   REGION "PAGE UP"
       //#hmi.page_up_actuate := #plc.pageUp.actuate;
       #hmi.page_up_animate := #plc.pageUp.animate;
       #hmi.page_up_enable := #plc.pageUp.enable;
       #hmi.page_up_label := #plc.pageUp.label;
       #hmi.page_up_list_select := #plc.pageUp.listSelect;
       #hmi.page_up_visible := #plc.pageUp.visible;
   END_REGION


   REGION "LINE UP"
       //#hmi.line_up_actuate := #plc.lineUp.actuate;
       #hmi.line_up_animate := #plc.lineUp.animate;
       #hmi.line_up_enable := #plc.lineUp.enable;
       #hmi.line_up_label := #plc.lineUp.label;
       #hmi.line_up_list_select := #plc.lineUp.listSelect;
       #hmi.line_up_visible := #plc.lineUp.visible;
   END_REGION


   REGION "LINE DOWN"
       //#hmi.line_down_actuate := #plc.lineDown.actuate;
       #hmi.line_down_animate := #plc.lineDown.animate;
       #hmi.line_down_enable := #plc.lineDown.enable;
       #hmi.line_down_label := #plc.lineDown.label;
       #hmi.line_down_list_select := #plc.lineDown.listSelect;
       #hmi.line_down_visible := #plc.lineDown.visible;
   END_REGION


   REGION "PAGE DOWN"
       //#hmi.page_down_actuate := #plc.pageDown.actuate;
       #hmi.page_down_animate := #plc.pageDown.animate;
       #hmi.page_down_enable := #plc.pageDown.enable;
       #hmi.page_down_label := #plc.pageDown.label;
       #hmi.page_down_list_select := #plc.pageDown.listSelect;
       #hmi.page_down_visible := #plc.pageDown.visible;
   END_REGION

   REGION "BOTTOM"
       //#hmi.bottom_actuate := #plc.bottom.actuate;
       #hmi.bottom_animate := #plc.bottom.animate;
       #hmi.bottom_enable := #plc.bottom.enable;
       #hmi.bottom_label := #plc.bottom.label;
       #hmi.bottom_list_select := #plc.bottom.listSelect;
       #hmi.bottom_visible := #plc.bottom.visible;
   END_REGION
END_FUNCTION

FUNCTION "NavBar: Private: First Row" : DInt   // FC180, SCL
{ S7_Optimized_Access := 'TRUE' }
VERSION : 0.1
   VAR_INPUT
      first_row : DInt;
      offset : DInt;
      TABLE_LENGTH : DInt;
   END_VAR
   VAR_TEMP
      ret : DInt;
   END_VAR
BEGIN
   REGION "DESCRIPTION"
       (*
       The new first row of the table is calculated from the offset. 
       Rollover and rollunder are resolved for the first row.
       *)
   END_REGION

   REGION "COPY TO INTERNAL"
       #ret := #first_row + #offset;
   END_REGION

   REGION "ROLLUNDER"
       IF #ret < 0 THEN
           #ret := #ret + #TABLE_LENGTH + 1;
       END_IF;
   END_REGION

   REGION "ROLLOVER"
       IF #ret > #TABLE_LENGTH THEN
           #ret := #ret - #TABLE_LENGTH - 1;
       END_IF;
   END_REGION

   REGION "OUTPUT"
       #"NavBar: Private: First Row" := #ret;
   END_REGION
END_FUNCTION

// folder: Utilities/Part Number

FUNCTION_BLOCK "IO Field: State Changes"   // FB48, SCL
{ S7_Optimized_Access := 'TRUE' }
VERSION : 0.1
   VAR_IN_OUT
      interface : "IO Field Data: Label with Data";
      feedback : "IO Field: State Change Data";
   END_VAR
   VAR
      old : "IO Field Data: Label with Data";
   END_VAR
BEGIN
   REGION "ANIMATE"
       #feedback.animate.rising := "USInt.Value_Change"(value := #interface.animate,
                                                         old_value := #old.animate);
       #feedback.animate.actual := #interface.animate;
       #feedback.animate.falling := FALSE;     // animate never set to null token 
   END_REGION

   REGION "ENABLE"
       #feedback.enable.rising := "Bool.Rising_Edge"(signal := #interface.enable,
                                                      old_signal := #old.enable);
       #feedback.enable.actual := #interface.enable;
       #feedback.enable.falling := "Bool.Falling_Edge"(signal := #interface.enable,
                                                        old_signal := #old.enable);
   END_REGION

   REGION "INPUT FINISHED"
       #feedback.input_finished.rising := "Bool.Rising_Edge"(signal := #interface.input_finished,
                                                              old_signal := #old.input_finished);
       #feedback.input_finished.actual := #interface.input_finished;
       #feedback.input_finished.falling := "Bool.Falling_Edge"(signal := #interface.input_finished,
                                                                old_signal := #old.input_finished);
   END_REGION

   REGION "VALUE CHANGED"
       #feedback.value.rising := "WString.Rising_Edge"(value := #interface.value,
                                                        old_value := #old.value);
       #feedback.value.actual := #interface.value;
       #feedback.value.falling := "WString.Falling_Edge"(value := #interface.value,
                                                          old_value := #old.value);
   END_REGION

   REGION "VISIBLE"
       #feedback.visible.rising := "Bool.Rising_Edge"(signal := #interface.visible,
                                                       old_signal := #old.visible);
       #feedback.visible.actual := #interface.visible;
       #feedback.visible.falling := "Bool.Falling_Edge"(signal := #interface.visible,
                                                         old_signal := #old.visible);
   END_REGION

   REGION "SAVE OLD VALUES"
       #old := #interface;
   END_REGION
END_FUNCTION_BLOCK

FUNCTION "Part_Number.Parse_Code" : Void   // FC34, SCL
{ S7_Optimized_Access := 'TRUE' }
VERSION : 0.1
   VAR_INPUT
      code : DInt;
   END_VAR
   VAR_OUTPUT
      code_left : DInt;
      code_right : DInt;
   END_VAR
BEGIN
   IF #code > 0 THEN
       #code_left := #code / 1000;
       #code_right := #code - #code / 1000 * 1000;
   ELSE
       #code_left := 0;
       #code_right := 0;
   END_IF;
END_FUNCTION

FUNCTION "Part_Number.Code_to_WString" : WString   // FC37, SCL
{ S7_Optimized_Access := 'TRUE' }
VERSION : 0.1
   VAR_INPUT
      pnLib : "Recipe: PN Text Library";
      pnCode : DInt;
   END_VAR
   VAR_TEMP
      pnLeft : DInt;
      pnRight : DInt;
      output : WString;
   END_VAR
   VAR CONSTANT
      newLine : WString := WSTRING#'$L';
   END_VAR
BEGIN
   REGION "PARSE CODE"
       "Part_Number.Parse_Code"(code := #pnCode,
                                 code_left => #pnLeft,
                                 code_right => #pnRight);
   END_REGION

   REGION "SINGLE LINE PN"
       IF "Part_Number.Is_Single"(#pnCode) THEN
           #output := #pnLib.pnText[#pnLeft];
       END_IF;
   END_REGION

   REGION "DOUBLE LINE PN"
       IF "Part_Number.Is_Double"(#pnCode) THEN
           #output := CONCAT_WSTRING(IN1 := #pnLib.pnText[#pnLeft],
                                     IN2 := #newLine,
                                     IN3 := #pnLib.pnText[#pnRight]);
       END_IF;
   END_REGION

   REGION "OUTPUT"
       #"Part_Number.Code_to_WString" := #output;
   END_REGION
END_FUNCTION

FUNCTION "Part_Number.Is_Double" : Bool   // FC153, SCL
{ S7_Optimized_Access := 'TRUE' }
VERSION : 0.1
   VAR_INPUT
      code : DInt;
   END_VAR
   VAR_TEMP
      code_left : DInt;
      code_right : DInt;
      ret : Bool;
   END_VAR
BEGIN
   REGION "NOTES"
       (*
       Double codes have a non-zero right hand component.
       Structure: XXXYYY
       XXX: left code, used for single and double codes
       YYY: right code, only used for double codes
       Last Edit: 2021-10-07
       *)
   END_REGION

   REGION "PROCESS CODE"
       "Part_Number.Parse_Code"(code := #code,
                                code_left => #code_left,
                                code_right => #code_right);
   END_REGION

   REGION "CHECK FOR DOUBLE CODE"
       IF #code_right > 0 THEN
           #ret := TRUE;
       END_IF;
   END_REGION

   REGION "RETURN" 
       #"Part_Number.Is_Double" := #ret;
   END_REGION
END_FUNCTION

FUNCTION "Part_Number.Is_Single" : Bool   // FC154, SCL
{ S7_Optimized_Access := 'TRUE' }
VERSION : 0.1
   VAR_INPUT
      code : DInt;
   END_VAR
   VAR_TEMP
      code_left : DInt;
      code_right : DInt;
      ret : Bool;
   END_VAR
BEGIN
   REGION "NOTES"
       (*
       Double codes have a non-zero right hand component.
       Structure:
       XXXYYY
       XXX: left code, used for single and double codes
       YYY: right code, only used for double codes
       Last Edit: 2021-10-07
       *)
   END_REGION

   REGION "PROCESS CODE"
       "Part_Number.Parse_Code"(code := #code,
                                code_left => #code_left,
                                code_right => #code_right);
   END_REGION

   REGION "CHECK FOR DOUBLE CODE"
       IF #code_right = 0 THEN
           #ret := TRUE;
       END_IF;
   END_REGION

   REGION "RETURN" 
       #"Part_Number.Is_Single" := #ret;
   END_REGION
END_FUNCTION

FUNCTION "Part_Number.WString_to_Code" : DInt   // FC240, SCL
{ S7_Optimized_Access := 'TRUE' }
VERSION : 0.1
   VAR_INPUT
      part_number : WString;
   END_VAR
   VAR_IN_OUT
      pn_library : "Recipe: PN Text Library";
   END_VAR
   VAR_TEMP
      _in_library : Bool;
      _library_full : Bool;
      _part_numbers : Array[0..1] of WString;
      _partial_pn_code : DInt;
      _pn_count : Int;
      _pn_code : DInt;
   END_VAR
   VAR CONSTANT
      OUT_OF_MEMORY : DInt := 999;
   END_VAR
BEGIN
   REGION "DATA PREP""
       "Part_Number.Split_PNs"(part_number := #part_number,
                               part_numbers := #_part_numbers);
       #_pn_count := "Part_Number.Count_PNs"(#_part_numbers);
   END_REGION


   REGION "NO PART NUMBERS ENTERED"
       IF #_pn_count = 0 THEN
           #"Part_Number.WString_to_Code" := 0;
           RETURN;
       END_IF;
   END_REGION


   REGION "CHECK FIRST PN CODE"
       #_pn_code := "Part_Number_Library.Search"(pn_library := #pn_library,
                                                 search_term := #_part_numbers[0]);
       #_in_library := "Part_Number.In_Library"(#_pn_code);
       #_library_full := "Part_Number_Library.Is_Full"(#pn_library);
   END_REGION


   REGION "FIRST PN CODE IN LIBRARY"
       IF #_in_library THEN
           #_pn_code *= 1_000;
       END_IF;
   END_REGION


   REGION "FIRST PN NOT IN LIBRARY, NO SPACE"
       IF NOT #_in_library AND #_library_full THEN
           #_pn_code := #OUT_OF_MEMORY * 1_000;
       END_IF;
   END_REGION


   REGION "FIRST PN NOT IN LIBRARY, SPACE"
       IF NOT #_in_library AND NOT #_library_full THEN
           #_pn_code := 1_000 * "Part_Number_Library.Add_PN"(pn := #_part_numbers[0],
                                                             pn_library := #pn_library);
       END_IF;
   END_REGION


   REGION "RETURN SINGLE PN CODE"
       IF #_pn_count = 1 THEN
           #"Part_Number.WString_to_Code" := #_pn_code;
           RETURN;
       END_IF;
   END_REGION


   REGION "CHECK SECOND PN CODE"
       #_partial_pn_code := "Part_Number_Library.Search"(pn_library := #pn_library,
                                                         search_term := #_part_numbers[1]);
       #_in_library := "Part_Number.In_Library"(#_partial_pn_code);
       #_library_full := "Part_Number_Library.Is_Full"(#pn_library);
   END_REGION


   REGION "SECOND PN CODE IN LIBRARY"
       IF #_in_library THEN
           #"Part_Number.WString_to_Code" := #_pn_code + #_partial_pn_code;
           RETURN;
       END_IF;
   END_REGION


   REGION "SECOND PN NOT IN LIBRARY, NO SPACE"
       IF NOT #_in_library AND #_library_full THEN
           #"Part_Number.WString_to_Code" := #_pn_code + #OUT_OF_MEMORY;
           RETURN;
       END_IF;
   END_REGION


   REGION "SECOND PN NOT IN LIBRARY, SPACE"
       IF NOT #_in_library AND NOT #_library_full THEN
           #_pn_code += "Part_Number_Library.Add_PN"(pn := #_part_numbers[1],
                                                     pn_library := #pn_library);
           #"Part_Number.WString_to_Code" := #_pn_code;
           RETURN;
       END_IF;
   END_REGION


   #"Part_Number.WString_to_Code" := 0;
   RETURN;
END_FUNCTION

FUNCTION "Part_Number.Count_PNs" : Int   // FC252, SCL
{ S7_Optimized_Access := 'TRUE' }
VERSION : 0.1
   VAR_INPUT
      part_numbers : Array[0..1] of WString;
   END_VAR
   VAR CONSTANT
      NULL : WString := WSTRING#'//';
      BLANK : WString := WSTRING#'';
   END_VAR
BEGIN
   IF #part_numbers[0] = #NULL THEN
       #"Part_Number.Count_PNs" := 0;
       RETURN;
   END_IF;

   IF #part_numbers[0] = #BLANK THEN
       #"Part_Number.Count_PNs" := 0;
       RETURN;
   END_IF;

   IF #part_numbers[1] = #NULL THEN
       #"Part_Number.Count_PNs" := 1;
       RETURN;
   END_IF;

   IF #part_numbers[1] = #BLANK THEN
       #"Part_Number.Count_PNs" := 1;
       RETURN;
   END_IF;

   #"Part_Number.Count_PNs" := 2;
   RETURN;
END_FUNCTION

FUNCTION "Part_Number.In_Library" : Bool   // FC253, SCL
{ S7_Optimized_Access := 'TRUE' }
VERSION : 0.1
   VAR_INPUT
      pn_code : DInt;
   END_VAR
BEGIN
   IF #pn_code = "NULL_TOKEN" THEN
       #"Part_Number.In_Library" := FALSE;
       RETURN;
   END_IF;
   #"Part_Number.In_Library" := TRUE;
   RETURN;
END_FUNCTION

FUNCTION "Part_Number.Split_PNs" : Void   // FC254, SCL
{ S7_Optimized_Access := 'TRUE' }
VERSION : 0.1
   VAR_INPUT
      part_number : WString;
   END_VAR
   VAR_IN_OUT
      part_numbers : Array[0..1] of WString;
   END_VAR
   VAR_TEMP
      _part_numbers : Array[0..1] of WString;
   END_VAR
   VAR CONSTANT
      NEW_LINE : WString := WSTRING#'$L';
      NULL : WString := WSTRING#'//';
   END_VAR
BEGIN
   "Array.WString.Fill"(value := #NULL,
                        array := #_part_numbers);
   "WString.Split_Single"(wstring_in := #part_number,
                          delimeter := #NEW_LINE,
                          "pointer" := 0,
                          sub_strings := #_part_numbers);
   #part_numbers := #_part_numbers;
END_FUNCTION

// folder: Utilities/Part Number Library

FUNCTION "Part_Number_Library.Is_Full" : Bool   // FC250, SCL
{ S7_Optimized_Access := 'TRUE' }
VERSION : 0.1
   VAR_INPUT
      pn_library : "Recipe: PN Text Library";
   END_VAR
   VAR_TEMP
      _first_null : DInt;
   END_VAR
   VAR CONSTANT
      NULL_STRING : WString := WSTRING#'//';
   END_VAR
BEGIN
   #_first_null := "Part_Number_Library.Search"(pn_library := #pn_library,
                                                search_term := #NULL_STRING);
   IF #_first_null = "NULL_TOKEN" THEN
       #"Part_Number_Library.Is_Full" := TRUE;
       RETURN;
   END_IF;

   #"Part_Number_Library.Is_Full" := FALSE;
   RETURN;
END_FUNCTION

FUNCTION "Part_Number_Library.Add_PN" : DInt   // FC251, SCL
{ S7_Optimized_Access := 'TRUE' }
VERSION : 0.1
   VAR_INPUT
      pn : WString;
   END_VAR
   VAR_IN_OUT
      pn_library : "Recipe: PN Text Library";
   END_VAR
   VAR_TEMP
      _index : DInt;
   END_VAR
   VAR CONSTANT
      NULL_STRING : WString := WSTRING#'//';
   END_VAR
BEGIN
   #_index := "Part_Number_Library.Search"(pn_library := #pn_library,
                                           search_term := #NULL_STRING);
   #pn_library.pnText[#_index] := #pn;
   #"Part_Number_Library.Add_PN" := #_index;
END_FUNCTION

FUNCTION "Part_Number_Library.Search" : Int   // FC255, SCL
{ S7_Optimized_Access := 'TRUE' }
VERSION : 0.1
   VAR_INPUT
      pn_library : "Recipe: PN Text Library";
      search_term : WString;
   END_VAR
   VAR_TEMP
      _array : Array[0..#MAX_ELEMENTS] of WString;
      _slices : Int;
      _slice : Int;
      _internal_length : Int;
      _external_length : Int;
      _search_result : Int;
   END_VAR
   VAR CONSTANT
      MAX_ELEMENTS : Int := 24;
   END_VAR
BEGIN
   REGION "NOTES"
       (*
           Why is this necessary?
               Unfortunately, dynamically sized arrays of wstring data type cannot accept
               wstrings of a declared length (e.x. the input parameter array[*] of 
               wstring[10] cannot exist). We need this wrapper function so that we can 
               copy wstrings of a declared length to an array of wstrings of default 
               length. Once copied, this array can be passed into the wstring search 
               function. However, there is only 16k of local memory to store the array of
               wstrings of default length. The pn text library can store up to 1000 part 
               numbers. If we were to copy all 1000, we would need 500k of memory. So, we 
               must slice the pn library into chunks and search them.
           Why are part number text wstrings a declared length?
               The declared lenght was necessary to fit a reasonable number of part 
               numbers into retentive memory.
       *)
   END_REGION


   REGION "SETUP"
       #_internal_length := UDINT_TO_INT("Array.Any.Length"(#_array));
       #_external_length := UDINT_TO_INT("Array.Any.Length"(#pn_library.pnText));
       #_slices := #_external_length / #_internal_length - 1;
   END_REGION


   REGION "REPEAT FOR EACH SLICE OF EXTERNAL ARRAY"
       FOR #_slice := 0 TO #_slices DO
           "Part_Number_Library.Search.Map_to_Internal_Array"(pn_library := #pn_library,
                                                              slice_number := #_slice,
                                                              internal_array := #_array);
           #_search_result := "Array.WString.Search"(array := #_array,
                                                     search_term := #search_term);
           IF #_search_result <> "NULL_TOKEN" THEN
               #"Part_Number_Library.Search" := #_search_result + #_slice * #_internal_length;
               RETURN;
           END_IF;
       END_FOR;
   END_REGION

   REGION "RETURN"
       #"Part_Number_Library.Search" := "NULL_TOKEN";
       RETURN;
   END_REGION
END_FUNCTION

FUNCTION "Part_Number_Library.Search.Map_to_Internal_Array" : Void   // FC256, SCL
{ S7_Optimized_Access := 'TRUE' }
VERSION : 0.1
   VAR_INPUT
      pn_library : "Recipe: PN Text Library";
      slice_number : Int;
   END_VAR
   VAR_IN_OUT
      internal_array : Array[*] of WString;
   END_VAR
   VAR_TEMP
      _i : Int;
      _length : Int;
      _p : Int;
   END_VAR
BEGIN
   #_length := UDINT_TO_INT("Array.Any.Length"(#internal_array));
   FOR #_i := 0 TO #_length - 1 DO
       #_p := #_i + #slice_number * #_length;
       #internal_array[#_i] := #pn_library.pnText[#_p];
   END_FOR;
END_FUNCTION

// folder: Utilities/Real

FUNCTION_BLOCK "Real.State_Change"   // FB52, SCL
{ S7_Optimized_Access := 'TRUE' }
VERSION : 0.1
   VAR_INPUT
      value : Real;
   END_VAR
   VAR_IN_OUT
      get_real : "State Changes: Real";
   END_VAR
   VAR
      old_value : Real;
   END_VAR
   VAR_TEMP
      _return : "State Changes: Real";
   END_VAR
BEGIN
   REGION "BUFFER IN"
       #_return := #get_real;
   END_REGION

   REGION "MAP"
       IF #value <> #old_value THEN
           #_return.actual := #value;
       END_IF;
       // these are set to false because there are no invalid times
       // negative should count in reverse
       // zero is valid
       #_return.rising := FALSE;
       #_return.falling := FALSE;
   END_REGION

   REGION "SAVE OLD VALUE"
       #old_value := #value;
   END_REGION


   REGION "RETURN" 
       #get_real := #_return;
   END_REGION
END_FUNCTION_BLOCK

// folder: Utilities/Screen Objects

FUNCTION "Cell_Data.Hide" : "Cell Data"   // FC209, SCL
{ S7_Optimized_Access := 'TRUE' }
VERSION : 0.1
BEGIN
   #"Cell_Data.Hide".animate := "INVISIBLE";
   #"Cell_Data.Hide".data := "BLANK";
   #"Cell_Data.Hide".visibility := "HIDE";
END_FUNCTION

FUNCTION "Cell_Data.Show" : "Cell Data"   // FC216, SCL
{ S7_Optimized_Access := 'TRUE' }
VERSION : 0.1
   VAR_INPUT
      animate : Int;
      data : WString;
   END_VAR
   VAR_TEMP
      _ret : "Cell Data";
   END_VAR
BEGIN
   #_ret.animate := #animate;
   #_ret.data := #data;
   #_ret.visibility := "SHOW";
   #"Cell_Data.Show" := #_ret;
END_FUNCTION

// folder: Utilities/Selected Buttons

FUNCTION "Selected_Buttons.Indices" : Void   // FC246, SCL
{ S7_Optimized_Access := 'TRUE' }
VERSION : 0.1
   VAR_INPUT
      selected_buttons : "Selected Buttons";
   END_VAR
   VAR_IN_OUT
      selected_buttons_indices : Array[*] of Int;
   END_VAR
   VAR_TEMP
      _i : Int;
      _length : Int;
      _resized_bool_array : Array[0..999] of Bool;
   END_VAR
BEGIN
   "Array.Bool.True_Indices"(array_of_bool := #selected_buttons.btns,
                             length := "BUTTON_COUNT",
                             list_of_indices := #selected_buttons_indices);
   FOR #_i := 0 TO "BUTTON_COUNT" DO
       IF #selected_buttons_indices[#_i] = "NULL_TOKEN" THEN
           CONTINUE;
       END_IF;
       #selected_buttons_indices[#_i] := "KP8.DURL_to_LRUD"(#selected_buttons_indices[#_i]);
   END_FOR;
END_FUNCTION

FUNCTION "Selected_Buttons.Get_First_Selected_Button" : Int   // FC289, SCL
{ S7_Optimized_Access := 'TRUE' }
VERSION : 0.1
   VAR_INPUT
      selected_buttons : "Selected Buttons";
   END_VAR
   VAR_TEMP
      _selected_buttons : Array[0.."BUTTON_COUNT"] of Int;
   END_VAR
BEGIN
   "Selected_Buttons.Indices"(selected_buttons := #selected_buttons,
                              selected_buttons_indices := #_selected_buttons);
   #"Selected_Buttons.Get_First_Selected_Button" := #_selected_buttons[0];
END_FUNCTION

// folder: Utilities/Selected Stations

FUNCTION "Selected_Stations.Indices" : Void   // FC245, SCL
{ S7_Optimized_Access := 'TRUE' }
VERSION : 0.1
   VAR_INPUT
      selected_stations : "Selected Stations";
   END_VAR
   VAR_IN_OUT
      selected_stations_indices : Array[*] of Int;
   END_VAR
   VAR_TEMP
      _i : Int;
      _length : Int;
      _resized_array : Array[0..999] of Bool;
   END_VAR
BEGIN
   FOR #_i := 0 TO "STATION_COUNT" DO
       #_resized_array[#_i] := #selected_stations.stns[#_i];
   END_FOR;
   "Array.Bool.True_Indices"(array_of_bool := #_resized_array,
                             length := "STATION_COUNT",
                             list_of_indices := #selected_stations_indices);
END_FUNCTION

FUNCTION "Selected_Stations.Matching_Line_Names" : Bool   // FC257, SCL
{ S7_Optimized_Access := 'TRUE' }
VERSION : 0.1
   VAR_INPUT
      stations : "Station: All Stations";
      selected_stations : "Selected Stations";
   END_VAR
   VAR_TEMP
      _i : Int;
      _first_selected_line_name : WString;
   END_VAR
   // Ret_Val : returns true when any number of stations selected and all selected stations have matching names
   VAR CONSTANT
      BLANK : WString;
   END_VAR
BEGIN
   REGION "NOTES"
       (*
           2022-04-06
           returns true if all selected stations have matching names
           returns false if no station selected
           returns false if selected stations do not have matching names
       *)
   END_REGION


   REGION "RETURN FALSE IF NO STATIONS SELECTED"
       IF #selected_stations.count = 0 THEN
           #"Selected_Stations.Matching_Line_Names" := FALSE;
           RETURN;
       END_IF;
   END_REGION


   REGION "CHECK EACH STATION"
       FOR #_i := 0 TO "STATION_COUNT" DO

           REGION "IGNORE DE-SELECTED STATIONS"
               IF NOT #selected_stations.stns[#_i] THEN
                   CONTINUE;
               END_IF;
           END_REGION

           REGION "SAVE FIRST SELECTED STATION'S NAME"
               IF #_first_selected_line_name = #BLANK THEN
                   #_first_selected_line_name := #stations.stn[#_i].id.lineName;
                   CONTINUE;
               END_IF;
           END_REGION

           REGION "RETURN FALSE IF SELECTED STATIONS' NAMES DO NOT MATCH"
               IF #_first_selected_line_name <> #stations.stn[#_i].id.lineName THEN
                   #"Selected_Stations.Matching_Line_Names" := FALSE;
                   RETURN;
               END_IF;
           END_REGION

       END_FOR;
   END_REGION


   REGION "ALL SELECTED STATIONS HAVE MATCHING NAMES"
       #"Selected_Stations.Matching_Line_Names" := TRUE;
   END_REGION
END_FUNCTION

FUNCTION "Selected_Stations.Get_First_Selected_Station" : Int   // FC274, SCL
{ S7_Optimized_Access := 'TRUE' }
VERSION : 0.1
   VAR_INPUT
      selected_stations : "Selected Stations";
   END_VAR
   VAR_TEMP
      _selected_stations : Array[0.."STATION_COUNT"] of Int;
   END_VAR
BEGIN
   "Selected_Stations.Indices"(selected_stations := #selected_stations,
                               selected_stations_indices := #_selected_stations);
   #"Selected_Stations.Get_First_Selected_Station" := #_selected_stations[0];
END_FUNCTION

// folder: Utilities/String

FUNCTION "Strip Sign" : WString   // FC3, SCL
{ S7_Optimized_Access := 'TRUE' }
VERSION : 0.1
   VAR_INPUT
      WString : WString;
   END_VAR
   VAR_TEMP
      Length : Int;
      "String Box" : WString;
      "Test Character" : WString;
   END_VAR
   VAR CONSTANT
      "+" : WChar := WCHAR#'+';
      "-" : WChar := WCHAR#'-';
   END_VAR
BEGIN
   #"String Box" := #WString;
   #"Test Character" := LEFT_WSTRING(IN := #"String Box",
                                     L := 1);
   IF #"Test Character" = #"+" OR #"Test Character" = #"-" THEN
       #Length := LEN(#"String Box");
       #"String Box" := RIGHT_WSTRING(IN := #"String Box", L := #Length - 1);

   END_IF;
   #"Strip Sign" := #"String Box";
END_FUNCTION

FUNCTION "Add Leading" : WString   // FC4, SCL
{ S7_Optimized_Access := 'TRUE' }
VERSION : 0.1
   VAR_INPUT
      "Leading Character" : WChar;
      "Desired Length" : USInt;
      "String" : WString;
   END_VAR
   VAR_TEMP
      Length : Int;
      "String Box" : WString;
   END_VAR
BEGIN
   #"String Box" := #String;
   #Length := LEN(#"String Box");

   WHILE #Length < #"Desired Length" DO
       #"String Box" := CONCAT_WSTRING(IN1 := #"Leading Character",
                                       IN2 := #"String Box");
       #Length := LEN(#"String Box");
   END_WHILE;

   #"Add Leading" := #"String Box";
END_FUNCTION

FUNCTION "WString.Word_Wrap_Depricated" : WString   // FC28, SCL
{ S7_Optimized_Access := 'TRUE' }
VERSION : 0.1
   VAR_INPUT
      stringIn : WString;
      maxLength : Int;
   END_VAR
   VAR_TEMP
      length : Int;
      lineBox : Array[0..#limitLines] of WString["LONG_STRING_LENGTH"];
      ret : WString;
      stringBox : Array[0..#limitString] of WString["LONG_STRING_LENGTH"];
   END_VAR
   VAR CONSTANT
      space : WString := WSTRING#' ';
      blank : WString;
      lineBreak : WString := WSTRING#'$L';
      limitString : Int := 49;
      limitLines : Int := 9;
   END_VAR
BEGIN
   REGION "GET LENGTH"
       #length := LEN(#stringIn);
   END_REGION

   REGION "NO WRAP NECESSARY"
       IF #length <= #maxLength THEN
           #ret := #stringIn;
       END_IF;
   END_REGION


   REGION "EXECUTE WORD WRAP"
       IF #length > #maxLength THEN

           "Explode"(stringIn := #stringIn,
                     explodedString := #stringBox);

           "WString.Word_Wrap_Depricated.Construct_Line"(stringBox := #stringBox,
                                       lineBox := #lineBox,
                                       maxLength := #maxLength);

           #ret := "WString.Word_Wrap_Depricated.Concat_Lines"(#lineBox);

       END_IF;
   END_REGION

   REGION "RETURN"
       #"WString.Word_Wrap_Depricated" := #ret;
   END_REGION
END_FUNCTION

FUNCTION "Trim" : WString   // FC29, SCL
{ S7_Optimized_Access := 'TRUE' }
VERSION : 0.1
   VAR_INPUT
      wString : WString;
   END_VAR
   VAR_TEMP
      ret : WString;
   END_VAR
   VAR CONSTANT
      space : WString := WSTRING#' ';
   END_VAR
BEGIN
   #ret := #wString;
   WHILE LEFT(IN := #ret, L := 1) = #space DO
       #ret := RIGHT(IN := #ret, L := LEN(#ret) - 1);
   END_WHILE;
   WHILE RIGHT(IN := #ret, L := 1) = #space DO
       #ret := LEFT(IN := #ret, L := LEN(#ret) - 1);
   END_WHILE;
   #Trim := #ret;
END_FUNCTION

FUNCTION "Upper" : Void   // FC49, SCL
{ S7_Optimized_Access := 'TRUE' }
VERSION : 0.1
   VAR_IN_OUT
      "string" : Variant;
   END_VAR
   VAR_TEMP
      "type" : Bool;
      stringBox : String;
      status : Int;
      wStringBox : WString;
      charArr : Array[0..255] of Char;
      cntChar : UInt;
      pChar : Int;
   END_VAR
   VAR CONSTANT
      asciiLow : Char := 'a';
      asciiHigh : Char := 'z';
      asciiCaseOffset : Int := 32;
   END_VAR
BEGIN
   IF TypeOf(#string) = String THEN
       #status := MOVE_BLK_VARIANT(SRC := #string,
                                   COUNT := 1,
                                   SRC_INDEX := 0,
                                   DEST_INDEX := 0,
                                   DEST => #stringBox);
   ELSIF TypeOf(#string) = WString THEN
       #status := MOVE_BLK_VARIANT(SRC := #string,
                                   COUNT := 1,
                                   SRC_INDEX := 0,
                                   DEST_INDEX := 0,
                                   DEST => #wStringBox);
       #stringBox := WSTRING_TO_STRING(#wStringBox);
   ELSE
       RETURN;
   END_IF;

   Strg_TO_Chars(Strg := #stringBox,
                 pChars := 0,
                 Cnt => #cntChar,
                 Chars := #charArr);

   FOR #pChar := 0 TO UINT_TO_INT(#cntChar) - 1 DO
       IF #asciiLow <= #charArr[#pChar] AND #charArr[#pChar] <= #asciiHigh THEN
           #charArr[#pChar] := INT_TO_CHAR(CHAR_TO_INT(#charArr[#pChar]) - #asciiCaseOffset);
       END_IF;
   END_FOR;

   Chars_TO_Strg(Chars := #charArr,
                 pChars := 0,
                 Cnt := #cntChar,
                 Strg => #stringBox);

   IF TypeOf(#string) = String THEN
       #status := MOVE_BLK_VARIANT(SRC := #stringBox,
                                   COUNT := 1,
                                   SRC_INDEX := 0,
                                   DEST_INDEX := 0,
                                   DEST => #string);
   ELSIF TypeOf(#string) = WString THEN
       #wStringBox := STRING_TO_WSTRING(#stringBox);
       #status := MOVE_BLK_VARIANT(SRC := #wStringBox,
                                   COUNT := 1,
                                   SRC_INDEX := 0,
                                   DEST_INDEX := 0,
                                   DEST => #string);
   END_IF;
END_FUNCTION

FUNCTION "Explode" : Void   // FC73, SCL
{ S7_Optimized_Access := 'TRUE' }
VERSION : 0.1
   VAR_INPUT
      stringIn : WString;
   END_VAR
   VAR_IN_OUT
      explodedString : Variant;
   END_VAR
   VAR_TEMP
      charBox : Array[0..#lmtChar] of WChar;
      count : DInt;
      pChar : Int;
      pStringBox : Int;
      stringBox : Array[0..#lmtString] of WString["LONG_STRING_LENGTH"];
      status : DInt;
   END_VAR
   VAR CONSTANT
      space : WString := WSTRING#' ';
      blank : WString;
      lineBreak : WString := WSTRING#'$L';
      lmtString : Int := 49;
      lmtChar : Int := 999;
   END_VAR
BEGIN
   Strg_TO_Chars(Strg := #stringIn,
                 pChars := 0,
                 Cnt => #count,
                 Chars := #charBox);

   FOR #pChar := 0 TO #count DO

       IF #charBox[#pChar] = #space THEN
           IF #charBox[#pChar + 1] = #space THEN
               EXIT;
           END_IF;
       END_IF;

       IF #pChar = 0 THEN
           #stringBox[#pStringBox] := #charBox[#pChar];
       END_IF;

       IF #pChar >= 1 THEN
           #stringBox[#pStringBox] := CONCAT_WSTRING(IN1 := #stringBox[#pStringBox],
                                                     IN2 := #charBox[#pChar]);
       END_IF;

       IF #charBox[#pChar] = #space THEN
           #stringBox[#pStringBox] := "Trim"(#stringBox[#pStringBox]);
           #pStringBox := #pStringBox + 1;
       END_IF;

       IF #charBox[#pChar] = #lineBreak THEN
           #stringBox[#pStringBox] := LEFT(IN := #stringBox[#pStringBox],
                                           L := LEN(#stringBox[#pStringBox]) - 1);
           #pStringBox := #pStringBox + 1;
           #stringBox[#pStringBox] := #lineBreak;
           #pStringBox := #pStringBox + 1;
       END_IF;

   END_FOR;

   #status := MOVE_BLK_VARIANT(SRC := #stringBox,
                               COUNT := INT_TO_UDINT(#pStringBox)+1,
                               SRC_INDEX :=0,
                               DEST_INDEX := 0,
                               DEST => #explodedString);
END_FUNCTION

FUNCTION "WString.Word_Wrap_Depricated.Construct_Line" : Void   // FC74, SCL
{ S7_Optimized_Access := 'TRUE' }
VERSION : 0.1
   VAR_INPUT
      stringBox : Array[0..#limitString] of WString["LONG_STRING_LENGTH"];
      maxLength : Int;
   END_VAR
   VAR_IN_OUT
      lineBox : Array[0..#limitLines] of WString["LONG_STRING_LENGTH"];
   END_VAR
   VAR_TEMP
      _lineBox : Array[0..#limitLines] of WString["LONG_STRING_LENGTH"];
      pString : Int;
      pLineBox : Int;
      lengthTest : WString;
   END_VAR
   VAR CONSTANT
      space : WString := WSTRING#' ';
      blank : WString;
      lineBreak : WString := WSTRING#'$L';
      limitString : Int := 49;
      limitLines : Int := 9;
   END_VAR
BEGIN
   REGION "FOR EACH STRING IN STRING LIST"
       FOR #pString := 0 TO #limitString DO

           REGION "END OF STRING LIST"
               IF #stringBox[#pString] = #blank THEN
                   IF #stringBox[#pString + 1] = #blank THEN
                       #_lineBox[#pLineBox] := "Trim"(#_lineBox[#pLineBox]);
                       #lineBox := #_lineBox;
                       RETURN;
                   END_IF;
               END_IF;
           END_REGION

           REGION "ON NEW LINE CHARACTER"
               IF #stringBox[#pString] = #lineBreak THEN
                   #_lineBox[#pLineBox] := "Trim"(#_lineBox[#pLineBox]);
                   #pLineBox := #pLineBox + 1;
                   #_lineBox[#pLineBox] := #lineBreak;
                   #pLineBox := #pLineBox + 1;
               END_IF;
           END_REGION

           REGION "BUILD EACH LINE"
               IF #stringBox[#pString] <> #lineBreak THEN

                   REGION "FIRST ELEMENT EDGE CASE"
                       IF #pString = 0 THEN
                           #lengthTest := #stringBox[#pString];
                       END_IF;
                   END_REGION

                   REGION "BUILT TEST STRING"
                       IF #pString >= 1 THEN
                           #lengthTest := CONCAT_WSTRING(IN1 := #_lineBox[#pLineBox],
                                                         IN2 := #space,
                                                         IN3 := #stringBox[#pString]);
                       END_IF;
                   END_REGION

                   REGION "TEST STRING NOT TOO LONG"
                       IF LEN(#lengthTest) <= #maxLength THEN
                           #_lineBox[#pLineBox] := #lengthTest;
                       END_IF;
                   END_REGION

                   REGION "TEST STRING TOO LONG"
                       IF LEN(#lengthTest) > #maxLength THEN
                           #_lineBox[#pLineBox] := "Trim"(#_lineBox[#pLineBox]);
                           #_lineBox[#pLineBox] := "Trim"(#_lineBox[#pLineBox]);
                           #pLineBox := #pLineBox + 1;
                           #_lineBox[#pLineBox] := #stringBox[#pString];
                       END_IF;
                   END_REGION

               END_IF;
           END_REGION

       END_FOR;
   END_REGION

   REGION "RETURN"
       #lineBox := #_lineBox;
   END_REGION
END_FUNCTION

FUNCTION "WString.Word_Wrap_Depricated.Concat_Lines" : WString   // FC75, SCL
{ S7_Optimized_Access := 'TRUE' }
VERSION : 0.1
   VAR_INPUT
      lineBox : Array[0..#limitLines] of WString["LONG_STRING_LENGTH"];
   END_VAR
   VAR_TEMP
      pLine : Int;
      ret : WString;
   END_VAR
   VAR CONSTANT
      space : WString := WSTRING#' ';
      blank : WString;
      lineBreak : WString := WSTRING#'$L';
      limitString : Int := 49;
      limitLines : Int := 9;
   END_VAR
BEGIN
   REGION "FOR EACH LINE"
       FOR #pLine := 0 TO #limitLines DO

           REGION "ON END OF LINE LIST"
               IF #lineBox[#pLine] = #space OR #lineBox[#pLine] = #blank THEN
                   EXIT;
               END_IF;
           END_REGION

           REGION "ON FIRST ELEMENT IN LINE LIST"
               IF #pLine = 0 THEN
                   #ret := #lineBox[#pLine];
               END_IF;
           END_REGION

           REGION "CONSTRUCT OUTPUT"
               IF #pLine >= 1 THEN

                   REGION "NO OP ON LINE BREAK CHARACTER"
                       IF #lineBox[#pLine] = #lineBreak THEN
                           ;// no action required
                       END_IF;
                   END_REGION

                   REGION "CONCATINATION"
                       IF #lineBox[#pLine] <> #lineBreak THEN
                           #ret := CONCAT_WSTRING(IN1 := #ret,
                                                  IN2 := #lineBreak,
                                                  IN3 := #lineBox[#pLine]);
                       END_IF;
                   END_REGION

               END_IF;
           END_REGION


       END_FOR;
   END_REGION

   REGION "RETURN"
       #ret := "Trim"(#ret);
       #"WString.Word_Wrap_Depricated.Concat_Lines" := #ret;
   END_REGION
END_FUNCTION

FUNCTION "WString.Split_Single" : Void   // FC202, SCL
{ S7_Optimized_Access := 'TRUE' }
VERSION : 0.1
   VAR_INPUT
      wstring_in : WString;
      delimeter : WString;
      pointer : Int;
   END_VAR
   VAR_IN_OUT
      sub_strings : Array[*] of WString;
   END_VAR
   VAR_TEMP
      _split : WString;
      _position : Int;
      _return : WString;
   END_VAR
BEGIN
   REGION "GET POSITION OF DELIMETER IN STRING"
       #_position := FIND(IN1 := #wstring_in,
                          IN2 := #delimeter);
   END_REGION

   REGION "BASE CASE"
       IF #_position = 0 THEN
           #sub_strings[#pointer] := #wstring_in;
           RETURN;
       END_IF;
   END_REGION


   REGION "RECURSIVE CASE"
       #sub_strings[#pointer] := LEFT(IN := #wstring_in, L := #_position - 1);
       "WString.Split_Single"(wstring_in := RIGHT(IN := #wstring_in, L := LEN(#wstring_in) - #_position),
                       delimeter := #delimeter,
                       "pointer" := #pointer + 1,
                       sub_strings := #sub_strings);
   END_REGION
END_FUNCTION

FUNCTION "WString.Word_Wrap" : WString   // FC203, SCL
{ S7_Optimized_Access := 'TRUE' }
VERSION : 0.1
   VAR_INPUT
      delimeters : Array[*] of WString[1];
      line_length : Int;
      wstring_in : WString;
   END_VAR
   VAR_TEMP
      _i : Int;
      _substring_length : Int;
      _wstring_in_length : Int;
      _pointer_substrings : Int;
      _substring : WString;
      _position_of_last_delimeter : Int;
      _recurse : Bool;
      _string_split_right : WString;
   END_VAR
   VAR CONSTANT
      BLANK : WString;
      NEW_LINE : WString := WSTRING#'$L';
   END_VAR
BEGIN
   #_wstring_in_length := LEN(#wstring_in);

   IF #line_length = 0 THEN
       #"WString.Word_Wrap" := #BLANK;
       RETURN;
   END_IF;

   FOR #_i := 1 TO #_wstring_in_length DO

       #_substring := CONCAT_WSTRING(IN1 := #_substring,
                                     IN2 := #wstring_in[#_i]);
       #_substring_length := LEN(#_substring);

       IF "Array.WString.Is_Element"(search_term := #wstring_in[#_i], search_array := #delimeters) THEN
           #_position_of_last_delimeter := #_i;
       END_IF;

       IF #wstring_in[#_i] = #NEW_LINE THEN
           #_substring := LEFT_WSTRING(IN := #_substring,
                                       L := #_substring_length - 1);
           #_string_split_right := RIGHT_WSTRING(IN := #wstring_in,
                                                 L := #_wstring_in_length - #_i);
           #_recurse := TRUE;
       END_IF;

       IF (#_substring_length = #line_length) AND (#_position_of_last_delimeter <> 0) THEN
           #_substring := LEFT_WSTRING(IN := #_substring,
                                       L := #_position_of_last_delimeter);
           #_string_split_right := RIGHT_WSTRING(IN := #wstring_in,
                                                 L := #_wstring_in_length - #_position_of_last_delimeter);
           #_recurse := TRUE;
       END_IF;

       IF (#_substring_length = #line_length) AND (#_position_of_last_delimeter = 0) THEN
           #_string_split_right := RIGHT_WSTRING(IN := #wstring_in,
                                                 L := #_wstring_in_length - #_substring_length);
           #_recurse := TRUE;
       END_IF;

       IF #_recurse THEN
           #_substring := CONCAT_WSTRING(IN1 := "Trim"(#_substring),
                                         IN2 := #NEW_LINE,
                                         IN3 := "WString.Word_Wrap"(delimeters := #delimeters,
                                                                    line_length := #line_length,
                                                                    wstring_in := #_string_split_right));
           #"WString.Word_Wrap" := #_substring;
           RETURN;
       END_IF;

   END_FOR; 

   #"WString.Word_Wrap" := "Trim"(#_substring);
END_FUNCTION

FUNCTION "WString.Find_Multiple.Depth" : Int   // FC204, SCL
{ S7_Optimized_Access := 'TRUE' }
VERSION : 0.1
   VAR_INPUT
      body : WString;
      terms : Array[*] of WString;
      p_terms : Int;
   END_VAR
   VAR_TEMP
      _length : UDInt;
      _position : Int;
   END_VAR
   VAR CONSTANT
      BLANK : WString;
   END_VAR
BEGIN
   (* 
       Depth first search of 'body' for first occurance of any element of 'terms'.
       For breadth first search, use WString.Find_Multiple.Breadth.
       Returns character postion in the string (1 indexed).
       E.G.: 
           - body := WSTRING#'today?'
           - terms := <WSTRING#>['?', 'ay']
           - returns --> 6
       E.G.:
           - body := WSTRING#'today?'
           - terms := <WSTRING#>['ay', '?']
           - returns --> 4
   *)

   #_length := "Array.Any.Length"(#terms);

   IF #p_terms > #_length OR #terms[#p_terms] = #BLANK THEN
           #"WString.Find_Multiple.Depth" := 0;
       RETURN;
   END_IF;

   #_position := FIND(IN1 := #body,
                      IN2 := #terms[#p_terms]);

   IF #_position = 0 THEN
       #_position := "WString.Find_Multiple.Depth"(body := #body,
                                             terms := #terms,
                                             p_terms := #p_terms + 1);
   END_IF;

   #"WString.Find_Multiple.Depth" := #_position;
END_FUNCTION

FUNCTION "WString.Find_Multiple.Breadth" : Int   // FC205, SCL
{ S7_Optimized_Access := 'TRUE' }
VERSION : 0.1
   VAR_INPUT
      body : WString;
      terms : Array[*] of WString[1];
   END_VAR
   VAR_TEMP
      _i : Int;
      _length : UDInt;
      _min : Int;
      _position : Int;
   END_VAR
   VAR CONSTANT
      BLANK : WString;
   END_VAR
BEGIN
   (* 
       Depth first search of 'body' for first occurance of any element of 'terms'.
       For depth first search use WString.Find_Multiple.Depth.
       Returns character postion in the string (1 indexed).
       E.G.: 
           - body := WSTRING#'today?'
           - terms := <WSTRING#>['?', 'ay']
           - returns --> 6
       E.G.:
           - body := WSTRING#'today?'
           - terms := <WSTRING#>['ay', '?']
           - returns --> 4
   *)

   #_length := "Array.Any.Length"(#terms);

   IF #_length = 0 OR #body = #BLANK THEN
       #"WString.Find_Multiple.Breadth" := 0;
       RETURN;
   END_IF;

   FOR #_i := 0 TO UDINT_TO_INT(#_length) - 1 DO
       #_position := FIND(IN1 := #body,
                          IN2 := #terms[#_i]);
       IF #_position = 0 THEN
           CONTINUE;
       END_IF;
       IF #_position < #_min OR #_min = 0 THEN
           #_min := #_position;
       END_IF;
   END_FOR;

   #"WString.Find_Multiple.Breadth" := #_min;
END_FUNCTION

FUNCTION "WString.Split_Multiple" : Void   // FC206, SCL
{ S7_Optimized_Access := 'TRUE' }
VERSION : 0.1
   VAR_INPUT
      wstring_in : WString;
      delimeters : Array[*] of WString[1];
      pointer : Int;
   END_VAR
   VAR_OUTPUT
      substrings : Array[*] of WString[20];
   END_VAR
   VAR_TEMP
      _i : Int;
      _position : Int;
      _return : WString;
      _split : WString;
   END_VAR
BEGIN
   REGION "GET POSITION OF DELIMETER IN STRING"
       #_position := "WString.Find_Multiple.Breadth"(body := #wstring_in,
                                                     terms := #delimeters);
   END_REGION

   REGION "BASE CASE"
       IF #_position = 0 THEN
           #substrings[#pointer] := #wstring_in;
           "WString.Split_Multiple.Clean_Output"("pointer" := #pointer + 1,
                                                 substrings := #substrings);
           RETURN;
       END_IF;
   END_REGION


   REGION "RECURSIVE CASE"
       #substrings[#pointer] := LEFT(IN := #wstring_in, L := #_position);
       "WString.Split_Multiple"(wstring_in := RIGHT(IN := #wstring_in, L := LEN(#wstring_in) - #_position),
                                delimeters := #delimeters,
                                "pointer" := #pointer + 1,
                                substrings => #substrings);
   END_REGION
END_FUNCTION

FUNCTION "WString.Split_Multiple.Clean_Output" : Void   // FC208, SCL
{ S7_Optimized_Access := 'TRUE' }
VERSION : 0.1
   VAR_INPUT
      pointer : Int;
   END_VAR
   VAR_IN_OUT
      substrings : Array[*] of WString;
   END_VAR
   VAR_TEMP
      _i : Int;
   END_VAR
   VAR CONSTANT
      BLANK : WString;
   END_VAR
BEGIN
   FOR #_i := #"pointer" TO UDINT_TO_INT("Array.Any.Length"(#substrings)) - 1 DO
       #substrings[#_i] := wstring#'';
   END_FOR;
END_FUNCTION

FUNCTION "Char.Is_Numeric" : Bool   // FC272, SCL
{ S7_Optimized_Access := 'TRUE' }
VERSION : 0.1
   VAR_INPUT
      character : Char;
   END_VAR
   VAR CONSTANT
      NUMBERS : String := '0123456789';
   END_VAR
BEGIN
   IF FIND(IN1 := #NUMBERS, IN2 := CHAR_TO_STRING(#character)) = 0 THEN
       #"Char.Is_Numeric" := FALSE;
       RETURN;
   END_IF;
   #"Char.Is_Numeric" := TRUE;
   RETURN;
END_FUNCTION

// folder: Utilities/Table Navigation

FUNCTION_BLOCK "Table Nav: End of Data Rollover"   // FB11, SCL
{ S7_Optimized_Access := 'TRUE' }
VERSION : 0.1
   VAR_INPUT
      tblData : Variant;
      tblDisp : Variant;
      nullFlag : Int;
      nullCheck : Variant;
      tableNav : "Nav Bar Data: PLC";
   END_VAR
   VAR_IN_OUT
      rowIndices : Variant;
   END_VAR
   VAR_TEMP
      firstNullIndex : DInt;
      len : Struct
         tblData : DInt;
         tblDisp : DInt;
      END_STRUCT;
      nullCheckVals : Array[0..#lenArrs] of DInt;
      offset : DInt;
      pulses : "Nav Bar Data: PLC";
      RET_VAL : Int;
      retRowIndices : Array[0..#lenArrs] of DInt;
   END_VAR
   VAR CONSTANT
      lenArrs : DInt := 999;
   END_VAR
BEGIN
       REGION "DESCRIPTION"
           (*
           Double checks row indicies against data and rolls over on end of data flag.
           *)
       END_REGION

       REGION "COPY TO LOCAL"
           #RET_VAL := MOVE_BLK_VARIANT(SRC := #rowIndices,
                                        COUNT := CountOfElements(#rowIndices),
                                        SRC_INDEX := 0,
                                        DEST_INDEX := 0,
                                        DEST => #retRowIndices);
           #RET_VAL := MOVE_BLK_VARIANT(SRC := #nullCheck,
                                        COUNT := CountOfElements(#nullCheck),
                                        SRC_INDEX := 0,
                                        DEST_INDEX := 0,
                                        DEST => #nullCheckVals);
       END_REGION

       REGION "GET ARRAY PARAMETERS"
           #len.tblData := UDINT_TO_DINT(CountOfElements(#tblData));
           #len.tblDisp := UDINT_TO_DINT(CountOfElements(#tblDisp));
       END_REGION

       REGION "CALCUALTE ROW INDICIES"
           "Table Nav: Calc Row Indices"(lenTblData := #firstNullIndex,
                                         lenTblDisp := #len.tblDisp,
                                         r1 := #retRowIndices[0],
                                         rowIndicies := #retRowIndices);
       END_REGION

       REGION "RETURN ROW INDICIES"
           #RET_VAL := MOVE_BLK_VARIANT(SRC := #retRowIndices,
                                        COUNT := DINT_TO_UDINT(#len.tblDisp),
                                        SRC_INDEX := 0,
                                        DEST_INDEX := 0,
                                        DEST => #rowIndices);
       END_REGION
END_FUNCTION_BLOCK

FUNCTION_BLOCK "Table Nav"   // FB43, SCL
{ S7_Optimized_Access := 'TRUE' }
VERSION : 0.1
   VAR_INPUT
      first_null_index : DInt;   // if you want to roll over before the end of your array, find the first null index and enter it here
      tblData : Variant;   // array to scan
      tblDisp : Variant;   // viewport array
      tableNav : "Nav Bar Data: PLC";   // table navigation udt
   END_VAR
   VAR_IN_OUT
      rowIndices : Variant;
   END_VAR
   VAR
      "inst Pulses: Table Nav" : "Table Nav: Pulses";
      r1 : DInt;
   END_VAR
   VAR_TEMP
      len : Struct
         tblData : DInt;
         tblDisp : DInt;
      END_STRUCT;
      offset : DInt;
      pulses : "Nav Bar Data: PLC";
      RET_VAL : Int;
      ret_row_indices : Array[0..#lenArrs] of DInt;
      ubound : DInt;
   END_VAR
   VAR CONSTANT
      lenArrs : DInt := 999;
   END_VAR
BEGIN
   REGION "DESCRIPTION"
       (*
       The function returns row indicies indicating the visible rows of a larger
       table determined by standard table navigation buttons.
       The function uses the variant data type to handle tables of any size.
       Rollover and rollunder features are built in.
       Row indices must be output to an array of dint (dimension is flexible).
       *)
   END_REGION


   REGION "GET PRESS PULSES"    
       #"inst Pulses: Table Nav"(press := #tableNav,
                                 pulses => #pulses);
   END_REGION


   REGION "RUN ON BUTTON PRESS"
       IF "Table Nav: Run Trigger"(#pulses) THEN